REGION Network 8: Störungsgruppe 2 und Änderung ermitteln; Bits -> DB für Anzeige
         L     4;  // Interner Offset für Störungsgruppe 2
         SLD   3;  // Anzahl der Bytes für die StGrp 1
         LAR1;  // Adresse für lokale Störungen
   //
         L     4;  // Interner Offset für Störungsgruppe 2
         L     #IN_Start_Stoerungen;
         +D;
         SLD   3;  //
         LAR2;  // Adresse für Störung im DB
   //
         L     1;  // Anzahl der Störungsworte
   M004: T     #Schleifenzaehler;  // Wenn Schleifenzähler <> 0
   //
         OPN   #IN_DB_Stoerungen;  //
         L     DBW[AR2, P#0.0];  // Gespeicherte Störung mit
         L     LW[AR1, P#0.0];  // Lokale Störung       vergleichen
         <>D;  //
         T     DBW[AR2, P#0.0];  // im DB speichern und
         S     #IO_Daten_Senden;  // Sendeanforderung an PU (FB120)
         S     #IO_Stoerungsaenderung;  // Störungsanderung für Störauswertung (FB9)
         S     #IO_Stoer_Grp_2_aktiv;  // und Sammelsignal setzen
   //
         +AR1  P#2.0;
         +AR2  P#2.0;
   //
         L     #Schleifenzaehler;  // Wenn Schleifenzähler <> 0
         LOOP  M004;  // Schleife erneut durchlaufen
   //
         A     #IN_Stoer_Grp_2_von_Ext;  // Störung vom Rechner
         AN    #IN_Reset_fault_Grp;  // in die SPS einbinden
         FP    #IO_FM_Stoer_Grp_2_v_Ext;
         S     #IO_Stoerungsaenderung;
         S     #IO_Stoer_Grp_2_aktiv;
END_REGION

REGION Network 9: Störungsgruppe 3 und Änderung ermitteln; Bits -> DB für Anzeige
         L     6;  // Interner Offset für Störungsgruppe 3
         SLD   3;  // Anzahl der Bytes für die StGrp 1 +2
         LAR1;  // Adresse für lokale Störungen
   //
         L     6;  // Interner Offset für Störungsgruppe 3
         L     #IN_Start_Stoerungen;
         +D;
         SLD   3;  //
         LAR2;  // Adresse für Störung im DB
   //
         L     3;  // Anzahl der Störungsworte
   M005: T     #Schleifenzaehler;  //
   //
         OPN   #IN_DB_Stoerungen;  //
         L     DBW[AR2, P#0.0];  // Gespeicherte Störung mit
         L     LW[AR1, P#0.0];  // Lokale Störung       vergleichen
         <>D;  //
         T     DBW[AR2, P#0.0];  // im DB speichern und
         S     #IO_Daten_Senden;  // Sendeanforderung an PU (FB120)
         S     #IO_Stoerungsaenderung;  // Störungsanderung für Störauswertung (FB9)
         S     #IO_Stoer_Grp_3_aktiv;  // und Sammelsignal setzen
   //
         +AR1  P#2.0;
         +AR2  P#2.0;
   //
         L     #Schleifenzaehler;  // Wenn Schleifenzähler <> 0
         LOOP  M005;  // Schleife erneut durchlaufen
   //
         A     #IN_Stoer_Grp_3_von_Ext;  // Storung vom Rechner
         AN    #IN_Reset_fault_Grp;  // in die SPS einbinden
         FP    #IO_FM_Stoer_Grp_3_v_Ext;
         S     #IO_Stoerungsaenderung;
         S     #IO_Stoer_Grp_3_aktiv;
END_REGION

REGION Network 10: Meldungen und Änderung ermitteln; Bits -> DB für Anzeige
         L     12;  // Interner Offset für Meldungen
         SLD   3;  //
         LAR1;  // Adresse für lokale Störungen
   //
         L     12;  // Interner Offset für Meldungen
         L     #IN_Start_Stoerungen;
         +D;
         SLD   3;  //
         LAR2;  // Adresse für Störung im DB
   //
         L     2;  // Anzahl der Meldungsworte
   M007: T     #Schleifenzaehler;  //
   //
         OPN   #IN_DB_Stoerungen;  //
         L     DBW[AR2, P#0.0];  // Gespeicherte Störung mit
         L     LW[AR1, P#0.0];  // Lokale Störung       vergleichen
         <>D;  //
         T     DBW[AR2, P#0.0];  // im DB speichern und
         S     #IO_Daten_Senden;  // Sendeanforderung an PU (FB120)
   //
         +AR1  P#2.0;
         +AR2  P#2.0;
   //
         L     #Schleifenzaehler;  // Wenn Schleifenzähler <> 0
         LOOP  M007;  // Schleife erneut durchlaufen
END_REGION
END_FUNCTION

FUNCTION "FC1019_Stoerauswertung" : Void   // FC1019, STL
TITLE = Stoerungsquittierung für 1 Formträger
{ S7_Optimized_Access := 'FALSE' }
AUTHOR : KT242
VERSION : 0.1
// Die Stoerungsquittierung erfolgt in zwei SPS-Zyklen: 
// 1.: mit Reset_fault_Fkt werden die Störungsbits der einzelnen FCs zurückgesetzt
// 2.: mit Reset_fault_Grp werden die Störungsbits der FCs für die Störungsgruppen
//     zurückgesetzt. Bilden diese nun die Störungen neu, so werten sie von
//     den einzelnen FCs bereits den aktuellen Stand aus, da diese bereits einen
//     SPS-Zyklus früher bearbeitet wurden.
// 
// Das Ablöschen der Störungen in der Visualisierung wird von den einzelnen 
// Stör-FCs organisiert.
   VAR_INPUT
      IN_Stoer_Grp_1_aktiv_RT : Bool;   // Störungsmerker für eine aktive Störung der Gruppe 1 an dem Rundtisch
      IN_Stoer_Grp_2_aktiv_RT : Bool;   // Störungsmerker für eine aktive Störung der Gruppe 2 an dem Rundtisch
      IN_Stoer_Grp_3_aktiv_RT : Bool;   // Störungsmerker für eine aktive Störung der Gruppe 3 an dem Rundtisch
      IN_Taster_Quittierung : Bool;   // Eingang für einen Taster zum quittieren der Störungen
      IN_Lampentest : Bool;   // Zur Überprüfung der Anzeigen wurde ein Lampentest angewählt
      IN_Erster_SPS_Zyklus : Bool;   // Impulssignal Neusstart der Steuerung zum ablöschen der Störungen
   END_VAR
   VAR_OUTPUT
      OUT_akustische_Anzeige : Bool;   // Ausgang für eine akustische Störungsanzeige (Nur bei Neustörungen)
      OUT_optische_Anzeige : Bool;   // Ausgang für eine optische Störungsanzeige
   END_VAR
   VAR_IN_OUT
      IO_Erste_Quittierung_oK : Bool;   // Hilfsmerker zum ablöschen der akustischen Störanzeige nach Quittierung
      IO_Reset_fault_Fkt : Bool;   // Signal zum quittieren der Störungen innerhalb der einzelnen Funktionsbausteine
      IO_Reset_fault_Grp : Bool;   // Signal zum quittieren der Störungen innerhalb der Störungsbausteine
      Stoerungsaenderung : Bool;   // Feststellen einer Störungsänderung für Abarbeitung
      IO_Quit_Flanke : Bool;   // Hilkfsmerker zur Überwachung der Betätigung des Quittiertasters
   END_VAR
   VAR_TEMP
      Sammel_Stoerung : Bool;   // Zwischenmerker für die erkennung einer anliegenden Störung
      Quit_Flanke : Bool;   // Zwischenmerker als Impuls für die Störungsquittierung
      Lampe_ein : Bool;   // Zwischenmerker für die Ansteuerung der optischen Störanzeige
   END_VAR
BEGIN

REGION Network 1: Störungsquittierung für die SPS
         NOP   0;
   //
   // Über das Bit Reset_fault_Fkt werden zuerst die Störungen
   // in den Funktionen in dem sie gebildet werden abgelöscht.
   // Im nächsten SPS- Zyklus werden dann erst die Störbits
   // in den jeweiligen Störungsbausteinen abgelöscht
   //
         A     #IO_Reset_fault_Grp;  // Für den Störungsbaustein
         R     #IO_Reset_fault_Grp;
   //
         A     #IO_Reset_fault_Fkt;  // Für die einzelnen Funktionsbausteine
         S     #IO_Reset_fault_Grp;
         R     #IO_Reset_fault_Fkt;
   //
   // Bilden einer Sammelstörung
   //
         O     #IN_Stoer_Grp_1_aktiv_RT;
         O     #IN_Stoer_Grp_2_aktiv_RT;
         O     #IN_Stoer_Grp_3_aktiv_RT;
         =     #Sammel_Stoerung;
   //
   // Quittierflanke gegen Dauerbetätigung des Quittiertasters
   //
         A     #IN_Taster_Quittierung;
         FP    #IO_Quit_Flanke;
         =     #Quit_Flanke;
   //
   // Wenn keine Störung mehr ansteht oder
   // wenn eine neue Störungsänderung erfolgt,
   // wird das Bit für die erste Quittierung zurückgesetzt
   //
         O     #Stoerungsaenderung;
         ON    #Sammel_Stoerung;
         R     #IO_Erste_Quittierung_oK;
   //
   // Wenn Störungen anstehen und zum 2´ten mal quittiert
   // wird wird das Quittierbit für die einzelnen FC´s
   // gesetzt
   //
         A     #Sammel_Stoerung;
         A     #IO_Erste_Quittierung_oK;
         A     #Quit_Flanke;
         S     #IO_Reset_fault_Fkt;
   //
   // Wurde die 2´te Quittierung an die einzelnen Maschinen
   // weitergegeben wird der Merker für die 1´te Quittierung
   // zurückgesetzt
   //
         A     #IO_Reset_fault_Fkt;
         R     #IO_Erste_Quittierung_oK;
   //
   // 1´tes mal quittieren -> Hupe ausschalten
   //
         A     #Sammel_Stoerung;
         AN    #Stoerungsaenderung;
         A     #Quit_Flanke;
         AN    #IO_Reset_fault_Fkt;
         S     #IO_Erste_Quittierung_oK;
   //
   // Störlampe immer wenn eine Störung ansteht
   //
         A     #Sammel_Stoerung;
         A     "Flag_01_000_Hertz";
         =     #Lampe_ein;
         O     #Lampe_ein;
         O     #IN_Lampentest;
         =     #OUT_optische_Anzeige;
   //
   // Störhupe nur wenn die erste Quittierung noch nicht erfolgte
   //
         O     #Lampe_ein;
         O     #IN_Lampentest;
         AN    #IO_Erste_Quittierung_oK;
         AN    #IN_Lampentest;
         =     #OUT_akustische_Anzeige;
   //
   // Bilden der Quittierungsbits zum ablöschen der einzelnen
   // Störungrn innerhalb der Funktionsbausteine
   //
         AN    #Sammel_Stoerung;
         A     #Quit_Flanke;
         O     #IN_Erster_SPS_Zyklus;  // Neustart der Steuerung
         S     #IO_Reset_fault_Fkt;
   //
   // Das Bit für die Anzeige einer Stoerungsaenderung
   // aus dem Störungsbaustein (FC1) wird zurücksetzen
   //
         SET;
         R     #Stoerungsaenderung;
END_REGION
END_FUNCTION

FUNCTION "FC1021_TT_Operation_mode" : Void   // FC1021, STL
TITLE = Betriebsarten der Anlage
{ S7_Optimized_Access := 'TRUE' }
VERSION : 0.1
   VAR_TEMP
      FRG_Start_Produktion : Bool;
      FRG_Produktion : Bool;
      FRG_Stop : Bool;
      Stopptaster : Bool;
      STG_GRP_2 : Bool;
      Temp_Auto_Stop_ok : Bool;
      Hupe_Anfahrwarnung : Bool;
      Anf_Stop : Bool;
   END_VAR
BEGIN

REGION Network 1
         A     "AS_turn_table";
         =     #Temp_Auto_Stop_ok;
         NOT;
         =     "DB1010_TT_Fault".AS.AS_Activ;
   //      =     "TT_H_AS"
END_REGION

REGION Network 2: Freigabesignale Produktion Starten bilden
         A     "DB1001_TT_State".BA_Anlage.Automatik_Stop_ok;
         A     "DB1001_TT_State".IPOS.Status.IPOS_referenziert;
         AN    "DB1001_TT_State".Bits.Stop_fuer_WW;
         AN    "DB1031_AddStatus".SaftyDevice[1].OpeningEnabled;
         AN    "DB1031_AddStatus".SaftyDevice[2].OpeningEnabled;
         AN    "DB1031_AddStatus".SaftyDevice[3].OpeningEnabled;
         AN    "DB1031_AddStatus".SaftyDevice[4].OpeningEnabled;
         =     #FRG_Start_Produktion;
END_REGION

REGION Network 3: Freigabesignale Produktionsbetrieb bilden
         A     "DB1001_TT_State".BA_Anlage.Start_Produktion;
         A     "DB1001_TT_State".IPOS.Status.RT_in_Position;
         =     #FRG_Produktion;
END_REGION

REGION Network 4: Freigabesignale Produktion Stoppen bilden
         A     "DB1001_TT_State".IPOS.Status.Stoppen_erkannt;
         A     "DB1001_TT_State".IPOS.Status.RT_in_Position;
         AN    "DB005_RS<->Extern".MC_Interface[1].Data_from_MC.Shot_preperation;
         =     #FRG_Stop;
END_REGION

REGION Network 5: Signal zum Stoppen bilden
         A     "Button_stop_cycle";
         AN    "DB1001_TT_State".Bits.Stop_fuer_WW;
         AN    "DB1001_TT_State".Bits.Stop_fuer_Teachen;
         AN    "DB1001_TT_State".Bits.StopAfterEmpty;
         A     "DB1001_TT_State".BA_Anlage.Automatik;
         =     #Stopptaster;
END_REGION

REGION Network 6: Bei Leerfahren der Anlage Störgruppe 2 ausblenden
         A     "DB1011_TT_Fault".STG2_RT;
         =     #STG_GRP_2;
END_REGION

REGION Network 7: Stoppen angefordert
         O     "DB1001_TT_State".Bits.Stop_fuer_WW;
         O     "DB1001_TT_State".Bits.Stop_fuer_Teachen;
         =     #Anf_Stop;
END_REGION

REGION Network 8: Funktion für Betriebsart
         CALL  "FC1022_TT_OM"
         ( IN_Steuerpannung        := "Controlvoltage_okay",
           IN_SS_Auto              := "Switch_automatic_mode",
           IN_SS_Hand              := "Switch_manual_mode",
           IN_Referenzieren        := "Button_reference_TT",
           IN_Automatik_Stop_ok    := #Temp_Auto_Stop_ok,
           IN_T_Start              := "Button_start_cycle",
           IN_T_Stop               := #Stopptaster,
           IN_Lampentest           := FALSE,
           IN_Werkzeugwechsel      := #Anf_Stop,
           IN_Freigabe_Start       := #FRG_Start_Produktion,
           IN_Freigabe_Produktion  := #FRG_Produktion,
           IN_Freigabe_Stop        := #FRG_Stop,
           IN_Stoerung_Gruppe_1    := "DB1011_TT_Fault".STG1_RT,
           IN_Stoerung_Gruppe_2    := #STG_GRP_2,
           IN_DW_Maxzeit_Prod_ein  := S5T#10S,
           IN_DW_Maxzeit_Prod_aus  := S5T#30S,
           IN_DW_Zeit_Startwarnung := "DB1049_TT_Value".Vorwarnzeit,
           IN_Betriebsart_Timer    := "TMTT_OPMode",
           IN_Anfahr_Timer         := "TMTT_StartProduction",
           IN_Produktions_Timer    := "TMTT_Production",
           Out_Anfahrwarnung       := #Hupe_Anfahrwarnung,
           IO_Status               := "DB1001_TT_State".BA_Anlage
         );
   //-----
END_REGION

REGION Network 9: Anzeige der Betriebsart der Anlage
         A     "DB1001_TT_State".BA_Anlage.Start_Produktion;
         A     "Flag_01_000_Hertz";
         O;
         A     "DB1001_TT_State".BA_Anlage.Produktion;
         A     "DB1001_TT_State".BA_Anlage.Stop_angefordert;
         A     "Flag_01_000_Hertz";
         O;
         A     "DB1001_TT_State".BA_Anlage.Produktion;
         AN    "DB1001_TT_State".BA_Anlage.Stop_angefordert;
         O     "DB1001_TT_State".BA_Anlage.Lampentest;
         =     "LED_start_cycle";
END_REGION

REGION Network 10: Leerfahren der Anlage ist beendet
   //      U     "T_Leerfahren_RT_1"
   //      FP    "FHM_RT_Leerfahren_RT1"
   //      =     "HM_RT_Leerfahren_RT1"
   //
   //      X     "HM_RT_Leerfahren_RT1"
   //      X     "DB005_RS<->Extern".Status_RT_1.S_RT_Leerfahren
   //      =     "DB005_RS<->Extern".Status_RT_1.S_RT_Leerfahren
   //
   //      U     #Starttaster
   //      R     "DB005_RS<->Extern".Status_RT_1.S_RT_Leerfahren
   // //
   //       U(
   //       O     "DB201_RT1_Segment_1".Status_FT.FT_aktuell.Status.FT_gesperrt
   //       O     "DB201_RT1_Segment_1".Status_FT.FT_aktuell.Status.FT_in_Abwahlposition
   //       )
   //       U(
   //       O     "DB202_RT1_Segment_2".Status_FT.FT_aktuell.Status.FT_gesperrt
   //       O     "DB202_RT1_Segment_2".Status_FT.FT_aktuell.Status.FT_in_Abwahlposition
   //       )
   //       U(
   //       O     "DB203_RT1_Segment_3".Status_FT.FT_aktuell.Status.FT_gesperrt
   //       O     "DB203_RT1_Segment_3".Status_FT.FT_aktuell.Status.FT_in_Abwahlposition
   //       )
   //       U(
   //       O     "DB204_RT1_Segment_4".Status_FT.FT_aktuell.Status.FT_gesperrt
   //       O     "DB204_RT1_Segment_4".Status_FT.FT_aktuell.Status.FT_in_Abwahlposition
   //       )
   //       U(
   //       O     "DB205_RT1_Segment_5".Status_FT.FT_aktuell.Status.FT_gesperrt
   //       O     "DB205_RT1_Segment_5".Status_FT.FT_aktuell.Status.FT_in_Abwahlposition
   //       )
   //       U(
   //       O     "DB206_RT1_Segment_6".Status_FT.FT_aktuell.Status.FT_gesperrt
   //       O     "DB206_RT1_Segment_6".Status_FT.FT_aktuell.Status.FT_in_Abwahlposition
   //       )
   //       U(
   //       O     "DB207_RT1_Segment_7".Status_FT.FT_aktuell.Status.FT_gesperrt
   //       O     "DB207_RT1_Segment_7".Status_FT.FT_aktuell.Status.FT_in_Abwahlposition
   //       )
   //       U(
   //       O     "DB208_RT1_Segment_8".Status_FT.FT_aktuell.Status.FT_gesperrt
   //       O     "DB208_RT1_Segment_8".Status_FT.FT_aktuell.Status.FT_in_Abwahlposition
   //       )
   //       U(
   //       O     "DB209_RT1_Segment_9".Status_FT.FT_aktuell.Status.FT_gesperrt
   //       O     "DB209_RT1_Segment_9".Status_FT.FT_aktuell.Status.FT_in_Abwahlposition
   //       )
   //       U(
   //       O     "DB210_RT1_Segment_10".Status_FT.FT_aktuell.Status.FT_gesperrt
   //       O     "DB210_RT1_Segment_10".Status_FT.FT_aktuell.Status.FT_in_Abwahlposition
   //       )
   //       U(
   //       O     "DB211_RT1_Segment_11".Status_FT.FT_aktuell.Status.FT_gesperrt
   //       O     "DB211_RT1_Segment_11".Status_FT.FT_aktuell.Status.FT_in_Abwahlposition
   //       )
   //       U(
   //       O     "DB212_RT1_Segment_12".Status_FT.FT_aktuell.Status.FT_gesperrt
   //       O     "DB212_RT1_Segment_12".Status_FT.FT_aktuell.Status.FT_in_Abwahlposition
   //       )
   //       U(
   //       O     "DB213_RT1_Segment_13".Status_FT.FT_aktuell.Status.FT_gesperrt
   //       O     "DB213_RT1_Segment_13".Status_FT.FT_aktuell.Status.FT_in_Abwahlposition
   //       )
   //       U(
   //       O     "DB214_RT1_Segment_14".Status_FT.FT_aktuell.Status.FT_gesperrt
   //       O     "DB214_RT1_Segment_14".Status_FT.FT_aktuell.Status.FT_in_Abwahlposition
   //       )
   //       U(
   //       O     "DB215_RT1_Segment_15".Status_FT.FT_aktuell.Status.FT_gesperrt
   //       O     "DB215_RT1_Segment_15".Status_FT.FT_aktuell.Status.FT_in_Abwahlposition
   //       )
   //       U(
   //       O     "DB216_RT1_Segment_16".Status_FT.FT_aktuell.Status.FT_gesperrt
   //       O     "DB216_RT1_Segment_16".Status_FT.FT_aktuell.Status.FT_in_Abwahlposition
   //       )
   //       U(
   //       O     "DB217_RT1_Segment_17".Status_FT.FT_aktuell.Status.FT_gesperrt
   //       O     "DB217_RT1_Segment_17".Status_FT.FT_aktuell.Status.FT_in_Abwahlposition
   //       )
   //       U(
   //       O     "DB218_RT1_Segment_18".Status_FT.FT_aktuell.Status.FT_gesperrt
   //       O     "DB218_RT1_Segment_18".Status_FT.FT_aktuell.Status.FT_in_Abwahlposition
   //       )
   //       U(
   //       O     "DB219_RT1_Segment_19".Status_FT.FT_aktuell.Status.FT_gesperrt
   //       O     "DB219_RT1_Segment_19".Status_FT.FT_aktuell.Status.FT_in_Abwahlposition
   //       )
   //       U(
   //       O     "DB220_RT1_Segment_20".Status_FT.FT_aktuell.Status.FT_gesperrt
   //       O     "DB220_RT1_Segment_20".Status_FT.FT_aktuell.Status.FT_in_Abwahlposition
   //       )
   //       =     "DB005_RS<->Extern".Status_RT_1.RT_ist_leergefahren
   // //
   //       U     "DB005_RS<->Extern".Status_RT_1.S_RT_Leerfahren
   //       UN    "DB005_RS<->Extern".Status_RT_1.RT_ist_leergefahren
   //       U     "Merker_01_000_Hertz"
   //       O(
   //       U     "DB005_RS<->Extern".Status_RT_1.RT_ist_leergefahren
   //       U     "DB005_RS<->Extern".Status_RT_1.S_RT_Leerfahren
   //       )
   //       O     "DB151_Rundtisch_1".BA_Anlage.Lampentest
   //       =     "H_Leerfahren_RT_1"
END_REGION
END_FUNCTION

FUNCTION "FC1022_TT_OM" : Void   // FC1022, STL
TITLE = Betriebsarten für die Anlage
{ S7_Optimized_Access := 'FALSE' }
AUTHOR : KT242
VERSION : 0.1
// Die Verwaltung der Betriebsarten geschieht wie folgt: 
// Die Betriebsarten hängen nur von der Stellung des Betriebsartenwahlschalters 
// ab, wie man es z.B. auch bei Robotern gewohnt ist. Das Bit "gültig" wurde in 
// "aktiv" geändert und zeigt zusätzlich, dass Steuerspannung und Schutztüren 
// o.k. sind.
// Referenzpunktfahren ist keine Betriebsart sondern ein zusätzliches Bit in 
// Betriebsart Hand.
// Automatikbetrieb hängt nicht davon ab, ob es möglich ist, die Anlage zu 
// bewegen. 
// Aggregate, die für den Automatikbetrieb nötig sind, sollten schon eingeschaltet 
// werden, wenn Betriebsart Automatik anliegt und Steuerspannung und NOTHALT o.k.
// sind.
   VAR_INPUT
      IN_Steuerpannung : Bool;   // Signal Steuerspannung Eingeschaltet und Not- Aus entriegelt
      IN_SS_Auto : Bool;   // Eingang Betriebsartenwahlschalter steht auf Automatik- Betrieb
      IN_SS_Hand : Bool;   // Eingang Betriebsartenwahlschalter steht auf Hand- Betrieb
      IN_Referenzieren : Bool;   // Eingang Taster für Referenzpunktfahrt
      IN_Automatik_Stop_ok : Bool;   // Eingang das die Sicherheitseinrichtungen quittiert sind
      IN_T_Start : Bool;   // Eingang für den Taster zum Starten des Rundtisches
      IN_T_Stop : Bool;   // Eingang für den Taster zum Stoppen des Rundtisches
      IN_Lampentest : Bool;   // Eingang für eine Funktionsüberprüfung der Lampenansteuerungen
      IN_Werkzeugwechsel : Bool;   // Signal das ein Werkzeugwechsel vorgewählt wurde
      IN_Freigabe_Start : Bool;   // Signal für die Freigabe zum Starten des Rundtisches
      IN_Freigabe_Produktion : Bool;   // Signal für die Freigabe des Produktionsbetriebes des Rundtisches
      IN_Freigabe_Stop : Bool;   // Signal für die Freigabe zum Stoppen des Rundtisches
      IN_Stoerung_Gruppe_1 : Bool;   // Eine Störung der Gruppe 1 steht an und wurde noch nicht quittiert
      IN_Stoerung_Gruppe_2 : Bool;   // Eine Störung der Gruppe 2 steht an und wurde noch nicht quittiert
      IN_DW_Maxzeit_Prod_ein : S5Time;   // Zeit in der die Produktion nach dem Starten freigegeben sein muß
      IN_DW_Maxzeit_Prod_aus : S5Time;   // Verzögerungszeit zum Stoppen des Produktionsbetriebes
      IN_DW_Zeit_Startwarnung : S5Time;   // Ansteuerungsdauer für eine Anfahrwarnung
      IN_Betriebsart_Timer : Timer;   // Timer für die Betriebsartenumschaltung
      IN_Anfahr_Timer : Timer;   // Timer für die Anfahrwarnung der Anlage
      IN_Produktions_Timer : Timer;   // Timer für die Produktions Start- und Abschaltung
   END_VAR
   VAR_OUTPUT
      Out_Anfahrwarnung : Bool;   // Ansteuerung einer Anfahrwarnung
   END_VAR
   VAR_IN_OUT
      IO_Status : "UDT_RT_Betriebsart";   // Speichern der Betriebsarten- Zustände für das Programm
   END_VAR
   VAR_TEMP
      Temp_IO_Status : "UDT_RT_Betriebsart";   // Temporärer Betriebsarten- Status für die interne Bearbeitung des Bausteins
      ERROR_CODE : Int;   // Störungszustand der Systemfunktion "BLKMOV" Blockmove
      Anyzeiger : ANY;   // Zeiger zum Kopieren der Bereiche "IO_Status" und "Temp_IO_Status"
      Ohne_Anfahrwarnung : Bool;   // Hilfsmerker das keine Anfahrwarnung benötigt wird
      Temp_Imp_Anfahrwarn_End : Bool;   // Impulsmerker das die Anfahrwarnung gerade beendet wurde
   END_VAR
BEGIN

REGION Network 1: Gesicherte Daten einbinden
         LAR1;
         L;
         LAR2;
   //
         L     W#16#1002;  // Bytes
         T     W[AR1, P#0.0];
         L     2;  // Anzahl Bytes
         T     W[AR1, P#2.0];
         L     W[AR2, P#0.0];  // Baustein Nr.
         T     W[AR1, P#4.0];
         L     D[AR2, P#2.0];  // Datenanfang
         T     D[AR1, P#6.0];
   //
         CALL  BLKMOV
         ( SRCBLK  := #Anyzeiger,
           RET_VAL := #ERROR_CODE,
           DSTBLK  := #Temp_IO_Status
         );
   //
END_REGION

REGION Network 2: Automatik- Stop
         A     #IN_Automatik_Stop_ok;
         =     #Temp_IO_Status.Automatik_Stop_ok;
END_REGION

REGION Network 3: Steuerspannung vorhanden
         A     #IO_Status.Steuerspannung_ein;
         JC    Spg;
   //
         A     #IN_Steuerpannung;
         L     S5T#1S;
         SD    #IN_Betriebsart_Timer;
         A     #IN_Betriebsart_Timer;
         =     #Temp_IO_Status.Steuerspannung_ein;
         JU    BA;
   //
   Spg:  A     #IN_Steuerpannung;
         =     #Temp_IO_Status.Steuerspannung_ein;
END_REGION

REGION Network 4: Wechsel der Betriebsart
         O(;
         AN    #IN_SS_Hand;
         A     #Temp_IO_Status.Hand;
         );
         O(;
         AN    #IN_SS_Auto;
         A     #Temp_IO_Status.Automatik;
         );
         L     S5T#500MS;
         SE    #IN_Betriebsart_Timer;
         A     #IN_Betriebsart_Timer;
         JC    GOON;
END_REGION

REGION Network 5: Betriebsartenschalter-Auswertung
   BA:   A     #IN_SS_Hand;
         AN    #IN_SS_Auto;
         =     #Temp_IO_Status.Hand;
   //
         AN    #IN_SS_Hand;
         A     #IN_SS_Auto;
         =     #Temp_IO_Status.Automatik;
   //
   GOON: A     #IN_Lampentest;
         =     #Temp_IO_Status.Lampentest;
   //
         O     #Temp_IO_Status.Hand;
         O     #Temp_IO_Status.Automatik;
         =     #Temp_IO_Status.Gueltig;
   //
         O     #Temp_IO_Status.Hand;
         O     #Temp_IO_Status.Automatik;
         A     #Temp_IO_Status.Steuerspannung_ein;
         A     #Temp_IO_Status.Automatik_Stop_ok;
         =     #Temp_IO_Status.Aktiv;
   //
         A     #Temp_IO_Status.Hand;
         A     #IN_Referenzieren;
         =     #Temp_IO_Status.Referenzieren;
END_REGION

REGION Network 6: Ausgabe eines Startsignales vor Ansteuerung der Anlage
         L     #IN_DW_Zeit_Startwarnung;
         L     0;
         ==D;
         =     #Ohne_Anfahrwarnung;
   //
         L     #IN_DW_Zeit_Startwarnung;
         A     #IN_Freigabe_Start;
         A     #IN_T_Start;
         A     #IN_T_Stop;
         A     #Temp_IO_Status.Automatik;
         AN    #IN_Stoerung_Gruppe_1;
         AN    #IN_Stoerung_Gruppe_2;
         AN    #Temp_IO_Status.Produktion;
         AN    #Temp_IO_Status.Start_Produktion;
         SE    #IN_Anfahr_Timer;
   //
         A     #IN_Anfahr_Timer;
         =     #Temp_IO_Status.Anfahrwarnung;
   //
         A     #Temp_IO_Status.Anfahrwarnung;
         =     #Out_Anfahrwarnung;
   //
         AN    #Temp_IO_Status.Anfahrwarnung;
         FP    #Temp_IO_Status.FHM_Anfahrwarnung;
         =     #Temp_Imp_Anfahrwarn_End;
END_REGION

REGION Network 7: Bit für Start Produktion
         L     #IN_DW_Maxzeit_Prod_ein;
         A     #IN_T_Start;
         A     #Ohne_Anfahrwarnung;
         O     #Temp_Imp_Anfahrwarn_End;
         A     #IN_Freigabe_Start;
         AN    #Temp_IO_Status.Produktion;
         AN    #Temp_IO_Status.Start_Produktion;
         S     #Temp_IO_Status.Start_Produktion;
         SE    #IN_Produktions_Timer;
   //
         ON    #IN_Produktions_Timer;
         ON    #Temp_IO_Status.Aktiv;
         ON    #Temp_IO_Status.Automatik;
         O     #IN_Stoerung_Gruppe_1;
         O     #IN_Stoerung_Gruppe_2;
         ON    #IN_T_Stop;
         O     #IN_Werkzeugwechsel;
         ON    #Temp_IO_Status.Automatik_Stop_ok;
         R     #Temp_IO_Status.Start_Produktion;
END_REGION

REGION Network 8: Bit für Produktion
         A     #Temp_IO_Status.Start_Produktion;
         A     #IN_Freigabe_Produktion;
         AN    #IN_Anfahr_Timer;
         S     #Temp_IO_Status.Produktion;
         R     #Temp_IO_Status.Start_Produktion;
   //
         L     #IN_DW_Maxzeit_Prod_aus;
         ON    #IN_T_Stop;
         O     #IN_Werkzeugwechsel;
         O     #IN_Stoerung_Gruppe_2;
         A     #Temp_IO_Status.Produktion;
         AN    #Temp_IO_Status.Stop_angefordert;
         S     #Temp_IO_Status.Stop_angefordert;
         SE    #IN_Produktions_Timer;
   //
         A     #Temp_IO_Status.Produktion;
         A     #IN_T_Start;
         AN    #IN_Werkzeugwechsel;
         R     #Temp_IO_Status.Stop_angefordert;
   //
         A     #Temp_IO_Status.Produktion;
         A     #Temp_IO_Status.Stop_angefordert;
         AN    #IN_Produktions_Timer;
         O;
         A     #Temp_IO_Status.Produktion;
         A     #Temp_IO_Status.Stop_angefordert;
         A     #IN_Freigabe_Stop;
         O     #IN_Stoerung_Gruppe_1;
         ON    #Temp_IO_Status.Automatik;
         ON    #Temp_IO_Status.Automatik_Stop_ok;
         ON    #Temp_IO_Status.Aktiv;
         R     #Temp_IO_Status.Produktion;
         R     #Temp_IO_Status.Stop_angefordert;
END_REGION

REGION Network 9: Daten sichern
         CALL  BLKMOV
         ( SRCBLK  := #Temp_IO_Status,
           RET_VAL := #ERROR_CODE,
           DSTBLK  := #Anyzeiger
         );
   //
END_REGION
END_FUNCTION

FUNCTION "FC1031_AdditionalDevice" : Void   // FC1031, STL
{ S7_Optimized_Access := 'TRUE' }
VERSION : 0.1
   VAR_TEMP
      Release_door : Bool;
      dummy : Bool;
   END_VAR
BEGIN

REGION Network 1: Safety door tool change
   //      UN    "DB1001_TT_State".BA_Anlage.Start_Produktion
   //      UN    "DB1001_TT_State".BA_Anlage.Produktion
   //      =     #Release_door
   //
   //      CALL  "FC1033_SafetyDevice"
   //         IN_With_Safety_door :=TRUE //"Settings_MCx".MC_settings.MCwithSafetydoor
   //         IN_EnableDoorOpen   :=#Release_door
   //         IN_SelectDoorOpen   :="Select_door_tool_change"
   //         IN_AS_Door          :="AS_door_tool_change"
   //         IN_QuitDoorOpen     :="Quit_door_tool_change"
   //         IN_OMLampTest       :="DB1001_TT_State".BA_Anlage.Lampentest
   //         IN_Delay_QuitDoor   :="TM_QuitDoor_MC1"
   //         OUT_V_DoorOpen      :="Release_door_tool_change"
   //         OUT_H_DoorOpen      :="Selected_door_tool_change"
   //         StatusSafetyDevice  :="DB1031_AddStatus".SaftyDevice[1]
END_REGION

REGION Network 2: Safety door robot
   //      UN    "DB1001_TT_State".BA_Anlage.Start_Produktion
   //      UN    "DB1001_TT_State".BA_Anlage.Produktion
   //      =     #Release_door
   //
   //      CALL  "FC1033_SafetyDevice"
   //         IN_With_Safety_door :=TRUE //"Settings_MCx".MC_settings.MCwithSafetydoor
   //         IN_EnableDoorOpen   :=#Release_door
   //         IN_SelectDoorOpen   :="Select_door_robot"
   //         IN_AS_Door          :="AS_door_robot"
   //         IN_QuitDoorOpen     :="Quit_door_robot"
   //         IN_OMLampTest       :="DB1001_TT_State".BA_Anlage.Lampentest
   //         IN_Delay_QuitDoor   :="TM_QuitDoor_MC1"
   //         OUT_V_DoorOpen      :="Release_door_robot"
   //         OUT_H_DoorOpen      :="Selected_door_robot"
   //         StatusSafetyDevice  :="DB1031_AddStatus".SaftyDevice[2]
END_REGION

REGION Network 3: Safety door test shot
END_REGION

REGION Network 4: Safety door turn table
   //      UN    "DB1001_TT_State".BA_Anlage.Start_Produktion
   //      UN    "DB1001_TT_State".BA_Anlage.Produktion
   //      =     #Release_door
   //
   //      CALL  "FC1033_SafetyDevice"
   //         IN_With_Safety_door :=TRUE //"Settings_MCx".MC_settings.MCwithSafetydoor
   //         IN_EnableDoorOpen   :=#Release_door
   //         IN_SelectDoorOpen   :="Select_door_TT"
   //         IN_AS_Door          :="AS_door_TT"
   //         IN_QuitDoorOpen     :="Quit_door_TT"
   //         IN_OMLampTest       :="DB1001_TT_State".BA_Anlage.Lampentest
   //         IN_Delay_QuitDoor   :="TM_QuitDoor_MC1"
   //         OUT_V_DoorOpen      :="Release_door_TT"
   //         OUT_H_DoorOpen      :="Selected_door_TT"
   //         StatusSafetyDevice  :="DB1031_AddStatus".SaftyDevice[3]

   //
END_REGION
END_FUNCTION

FUNCTION "FC1032_PneuZylindermSH" : Void   // FC1032, STL
TITLE = Pneumatischer Zylinder mit Selbsthaltung
{ S7_Optimized_Access := 'FALSE' }
VERSION : 0.1
   VAR_INPUT
      BA_Auto : Bool;   // Betriebsart Automatik
      BA_Hand : Bool;   // Tippbetrieb
      Anf_GS : Bool;   // Anforderung Grundstellung Automatik
      Anf_AS : Bool;   // Anforderung Arbeitsstellung Automatik
      T_GS : Bool;   // Taste Grundstellung (Tippbetrieb)
      T_AS : Bool;   // Taste Arbeitsstellung (Tippbetrieb)
      Frg_GS : Bool;   // Bewegungsbedingungen für Grundstellungsfahrt erfüllt
      Frg_AS : Bool;   // Bewegungsbedingungen für Arbeitstellungsfahrt erfüllt
      INI_GS : Bool;   // Sensorik Zylinder befindet sich in Grundstellung
      INI_AS : Bool;   // Sensorik Zylinder befindet sich in Arbeitsstellung
      P_GS : Bool;   // Druckschalter Grundstellung
      P_AS : Bool;   // Druckschalter Arbeitsstellung
      IN_Reset_fault_Fkt : Bool;   // Signal to acknowledge faults in functionblock
      Laufzeit : S5Time;   // Laufzeit für Laufzeitüberwachung
      TM_Laufzeit : Timer;   // Timer zur Laufzeitüberwachung
   END_VAR
   VAR_OUTPUT
      H_GS : Bool;   // Anzeige Grundstellung
      H_AS : Bool;   // Anzeige Arbeitsstellung
      OUT_V_GS : Bool;   // Ventil zur Ansteuerung der Grundstellung
      OUT_V_AS : Bool;   // Ventil zur Ansteuerung der Arbeitsstellung
   END_VAR
   VAR_IN_OUT
      IO_Stg_INI : Bool;   // Sensorstörung
      IO_Stg_Laufzeit : Bool;   // Laufzeitstörung
      IO_NewFault : Bool;
      IO_FaultLevel_1 : Bool;
   END_VAR
   VAR_TEMP
      Temp_V_GS : Bool;
      Temp_V_AS : Bool;
   END_VAR
BEGIN

REGION Network 1: Ausgänge Rücksetzen
         CLR;
         =     #Temp_V_GS;
         =     #Temp_V_AS;
END_REGION

REGION Network 2: Störungen zurücksetzen
         A     #IN_Reset_fault_Fkt;
         R     #IO_Stg_INI;
         R     #IO_Stg_Laufzeit;
END_REGION

REGION Network 3: Tippbetrieb
         A     #BA_Hand;
         JCN   nHnd;

   // Arbeitsstellung
         A     #T_AS;
         A     #Frg_AS;
         O(;
         A     #INI_AS;
         A     #P_AS;
         AN(;
         A     #T_GS;
         A     #Frg_GS;
         );
         );
         =     #Temp_V_AS;

   // Grundstellung
         A     #T_GS;
         A     #Frg_GS;
         O(;
         A     #INI_GS;
         A     #P_GS;
         AN(;
         A     #T_AS;
         A     #Frg_AS;
         );
         );
         =     #Temp_V_GS;

   nHnd: NOP   0;
END_REGION

REGION Network 4: Automatik
         A     #BA_Auto;
         JCN   nAut;

   // Arbeitsstellung
         A     #Anf_AS;
         A     #Frg_AS;
         O(;
         A     #INI_AS;
         A     #P_AS;
         AN(;
         A     #Anf_GS;
         A     #Frg_GS;
         );
         );
         =     #Temp_V_AS;

   // Grundstellung
         A     #Anf_GS;
         A     #Frg_GS;
         O(;
         A     #INI_GS;
         A     #P_GS;
         AN(;
         A     #Anf_AS;
         A     #Frg_AS;
         );
         );
         =     #Temp_V_GS;

   nAut: NOP   0;
END_REGION

REGION Network 5: Anzeigen

         A     #Temp_V_GS;
         =     #OUT_V_GS;
         A     #Temp_V_AS;
         =     #OUT_V_AS;

         ON    #INI_GS;
         ON    #P_GS;
         A     #Temp_V_GS;
         A     "Flag_01_250_Hertz";
         O(;
         A     #INI_GS;
         A     #P_GS;
         );
         =     #H_GS;

         ON    #INI_AS;
         ON    #P_AS;
         A     #Temp_V_AS;
         A     "Flag_01_250_Hertz";
         O(;
         A     #INI_AS;
         A     #P_AS;
         );
         =     #H_AS;
END_REGION

REGION Network 6: Störungen
   //  Sensorstörung
         A     #INI_GS;
         A     #INI_AS;
         AN    #IO_Stg_INI;
         S     #IO_NewFault;
         S     #IO_Stg_INI;

   //  Laufzeitstörung
         A(;

         O(;
         X     #Temp_V_GS;
         X(;
         A     #INI_GS;
         A     #P_GS;
         );
         );

         O(;
         X     #Temp_V_AS;
         X(;
         A     #INI_AS;
         A     #P_AS;
         );
         );
         );

         A(;
         O     #BA_Hand;
         O     #BA_Auto;
         );

         L     #Laufzeit;
         SD    #TM_Laufzeit;

         A     #TM_Laufzeit;
         AN    #IO_Stg_Laufzeit;
         S     #IO_NewFault;
         S     #IO_Stg_Laufzeit;
END_REGION
END_FUNCTION

FUNCTION "FC1033_SafetyDevice" : Void   // FC1033, STL
{ S7_Optimized_Access := 'FALSE' }
VERSION : 0.1
   VAR_INPUT
      IN_With_Safety_door : Bool;   // Input if safety door is available
      IN_EnableDoorOpen : Bool;   // Enable signal for the release to open the door
      IN_SelectDoorOpen : Bool;   // Input for the selection to open the door
      IN_AS_Door : Bool;   // Input from the saftey that the door is open
      IN_QuitDoorOpen : Bool;   // Input to reset the door clamping
      IN_OMLampTest : Bool;   // Operation mode for lamp test is selected
      IN_Delay_QuitDoor : Timer;
   END_VAR
   VAR_OUTPUT
      OUT_V_DoorOpen : Bool;   // Output valve to clamp the door
      OUT_H_DoorOpen : Bool;   // Output for the lamp
   END_VAR
   VAR_IN_OUT
      StatusSafetyDevice : "UDT_SafetyDevice";
   END_VAR
BEGIN

REGION Network 1: If deselect jump to delete
         A     #IN_With_Safety_door;
         JCN   delete;
END_REGION

REGION Network 2: Edge of the button to select opening of the safety device
   // Switch off delay for PILZ switch

         A     #IN_QuitDoorOpen;
         L     s5t#1s;
         SF    #IN_Delay_QuitDoor;
   //----
         A     #IN_SelectDoorOpen;
         FN    #StatusSafetyDevice.HFEdgeButton;
         =     #StatusSafetyDevice.EdgeButton;
   //----
         A     #IN_AS_Door;
         FP    #StatusSafetyDevice.HFEdgeASReset;
         =     #StatusSafetyDevice.EdgeASReset;
   //----
         X     #StatusSafetyDevice.EdgeButton;
         X     #StatusSafetyDevice.OpeningSelected;
         O     #StatusSafetyDevice.HFforMESAutomaticStop;
         AN    #StatusSafetyDevice.EdgeASReset;
         AN    #IN_Delay_QuitDoor;
         =     #StatusSafetyDevice.OpeningSelected;
   //----
         A     #StatusSafetyDevice.OpeningSelected;
         A     #IN_EnableDoorOpen;
   //      ON    #IN_Delay_QuitDoor
         =     #StatusSafetyDevice.OpeningEnabled;
         NOT;
         =     #OUT_V_DoorOpen;
   //----
         O     #StatusSafetyDevice.OpeningEnabled;
         O(;
         A     #StatusSafetyDevice.OpeningSelected;
         A     "Flag_01_000_Hertz";
         );
         ON    #IN_AS_Door;
         O     #IN_OMLampTest;
         =     #OUT_H_DoorOpen;
   //----
         A     #StatusSafetyDevice.OpeningSelected;
         =     #StatusSafetyDevice.HFforMESSelected;
   //----
         AN    #IN_AS_Door;
         =     #StatusSafetyDevice.HFforMESAutomaticStop;
         R     #StatusSafetyDevice.HFforMESSelected;
   //---
         A     #StatusSafetyDevice.HFforMESSelected;
         =     #StatusSafetyDevice.Msg_Selected;
         A     #StatusSafetyDevice.HFforMESAutomaticStop;
         =     #StatusSafetyDevice.Msg_AS_active;
   //---
         BEU;
END_REGION

REGION Network 3: Delete
   delete:SET;
         R     #StatusSafetyDevice.Msg_Selected;
         R     #StatusSafetyDevice.Msg_AS_active;
         R     #OUT_H_DoorOpen;
         R     #OUT_V_DoorOpen;
END_REGION
END_FUNCTION

FUNCTION "FC1040_TT_Movement" : Void   // FC1040, STL
TITLE = Ansteuern der Anlage
{ S7_Optimized_Access := 'TRUE' }
VERSION : 0.1
   VAR_TEMP
      Temp_Segmentinis : DWord;   // Hilfsmerker für die Positionserkennung über die Hardwareabschaltung im Zentrum
      Temp_Rampe_Plus : Int;   // Hilfswort für die Beschleunigung des Rundtisches
      Temp_Rampe_Minus : Int;   // Hilfswort für die Verzögerung des Rundtisches
      Temp_Speed_Hand : Int;   // Hilfswort für die Geschwindigkeit im Handbetrieb
      Temp_Speed_Automatik : Int;   // Hilfswort für die Geschwindigkeit im Automatikbetrieb
      Temp_Offset_Position : Int;   // Hilfswort für den negativen Offset bei einer Positionierung im kont. Betrieb
      Temp_AmoutOfSegments : Int;   // Help word to define the amount of segments
      Temp_Drehsperre : Bool;   // Hilfsmerker für die generelle Freigabe dere Anlage
      Temp_Taktfreigabe : Bool;   // Hilfsmerker für das Takten der Anlage
      Temp_Drehfreigabe : Bool;   // Hilfsmerker für die Freigabe zum Ansteuern der Anlage
      Temp_RT_in_Position : Bool;   // Hilfsmerker für die Umschaltung der Segmentpositionen
      Temp_GenauhalteSignal : Bool;   // Hilfsmerker für die Ermittlung des Genauhaltes
      Temp_AnfahrWarnung : Bool;   // Hilfsmerker für die Huppe als Anfahr Warnung
      Temp_AnfahrWarnung_1 : Bool;   // Hilfsmerker für die Huppe als Anfahr Warnung
   END_VAR
BEGIN

REGION Network 1: Amount of Segments
         L     4;
         T     #Temp_AmoutOfSegments;
END_REGION

REGION Network 2: Drehsperren auswerten
         A     "DB1001_TT_State".BA_Anlage.Automatik_Stop_ok;
   //      UN    "DB009_Faults".Faults_FKT_Grp_1_M1
         =     #Temp_Drehfreigabe;
         NOT;
         =     #Temp_Drehsperre;
END_REGION

REGION Network 3: Taktzeitverlängerung // Anlage anhalten
         A     "Button_extend_cycle";
         FP    "FHM_Takt_Verz_RT1";
         =     "HM_FP_Takt_Verz_RT1";

         A     "HM_FP_Takt_Verz_RT1";
         AN    "DB1001_TT_State".Bits.Taktdehnung;
         S     "DB1001_TT_State".Bits.Taktdehnung;
         JC    VERZ;

         A     "HM_FP_Takt_Verz_RT1";
         A     "DB1001_TT_State".Bits.Taktdehnung;
         R     "DB1001_TT_State".Bits.Taktdehnung;

   VERZ: NOP   0;
         ON    "DB1001_TT_State".BA_Anlage.Produktion;
         R     "DB1001_TT_State".Bits.Taktdehnung;
   //
         A     "DB1001_TT_State".Bits.Taktdehnung;
         AN    "DB1001_TT_State".IPOS.Status.RT_in_Position;
         A     "Flag_01_000_Hertz";
         O;
         A     "DB1001_TT_State".Bits.Taktdehnung;
         A     "DB1001_TT_State".IPOS.Status.RT_in_Position;
         A     "Flag_05_000_Hertz";
         O     "DB1001_TT_State".BA_Anlage.Lampentest;
         =     "LED_extend_cycle";
END_REGION

REGION Network 4: Freigabe zum Takten der Anlage

         AN    "DB1001_TT_State".Bits.Stop_fuer_WW;
         AN    "DB1001_TT_State".Bits.Stop_fuer_Teachen;
         AN    "DB1001_TT_State".Bits.StopAfterEmpty;

         AN    "DB005_RS<->Extern".MC_Interface[1].Data_from_MC.Shot_release;
         AN    "DB005_RS<->Extern".MC_Interface[1].Data_from_MC.Shot_preperation;
         AN    "DB1001_TT_State".BA_Anlage.Stop_angefordert;
         AN    "DB1030_TT_AddFaults".SafteyDeviceSelected[1];
         AN    "DB1030_TT_AddFaults".SafteyDeviceSelected[2];
         AN    "DB1030_TT_AddFaults".SafteyDeviceSelected[3];

         A     #Temp_Drehfreigabe;
         AN    "DB1001_TT_State".Bits.Taktdehnung;
         A     "DB1001_TT_State".BA_Anlage.Automatik;
         =     #Temp_Taktfreigabe;
END_REGION

REGION Network 5: Taktimpuls bilden
         CALL  "FC1041_TT_Taktimpuls"
         ( IN_Drehfreigabe         := #Temp_Taktfreigabe,
           IN_Taktfreigabe         := #Temp_Drehfreigabe,
           IN_Anlage_in_Position   := "DB1001_TT_State".IPOS.Status.RT_in_Position,
           IN_Start_Anlagenbetrieb := "DB1001_TT_State".BA_Anlage.Produktion,
           IN_Anlagenbetrieb       := "DB1001_TT_State".BA_Anlage.Start_Produktion,
           IN_DW_Taktzeit          := "DB1049_TT_Value".Taktzeit,
           IN_Takttimer            := "TMTT_Tact",
           IN_Vorwarnzeit_1_in_Dec := 5,
           IN_Vorwarnzeit_2_in_Dec := 3,
           IO_Status               := "DB1001_TT_State".Takt
         );
   //-----
END_REGION

REGION Network 6: Sollwerte an FU
         L     "DB1049_TT_Value".Antrieb_RP;
         T     #Temp_Rampe_Plus;
         L     "DB1049_TT_Value".Antrieb_RN;
         T     #Temp_Rampe_Minus;
         L     "DB1049_TT_Value".Antrieb_Hand;
         T     #Temp_Speed_Hand;
         L     "DB1049_TT_Value".Antrieb_Auto;
         T     #Temp_Speed_Automatik;
   //-----
         L     0;
         A     "DB1001_TT_State".Bits.Stop_fuer_WW;
         JCN   Off2;
         L     "DB1049_TT_Value".Pos_Offset_WW;
         JU    Off;
   Off2: NOP   0;
         A     "DB1001_TT_State".Bits.Stop_fuer_Teachen;
         JCN   Off3;
         L     "DB1049_TT_Value".Pos_Offset_Teachen;
         JU    Off;
   Off3: NOP   0;
   Off:  T     #Temp_Offset_Position;
END_REGION

REGION Network 7: Umrichter für Rundtisch ansteuern
         A     "Button_Tip_+";
         A     "DB1001_TT_State".BA_Anlage.Hand;
         =     "Button_Tip_+";

         A     "Button_Tip_-";
         A     "DB1001_TT_State".BA_Anlage.Hand;
         =     "Button_Tip_-";

   // Genauhalt INI
         L     "DB1001_TT_State".IPOS.Status.Aktuelle_Position;
         L     0;
         ==I;
         A     "DB1001_TT_State".IPOS.Eingaenge_von_IPOS.Ipos_referenziert;
         =     #Temp_GenauhalteSignal;
   //-----
         CALL  "FC1042_RT_IPOS_CTRL"
         ( IN_EA_Adresse            := 700,
           IN_Taktend               := TRUE,
           IN_Taktend_1_Segment     := TRUE,
           IN_DP_ok                 := TRUE,
           IN_IPOS_referenziert     := "DB1001_TT_State".IPOS.Eingaenge_von_IPOS.Ipos_referenziert,
           IN_Stoerung_Luefter      := FALSE,
           IN_Motorschutz           := "F_FC_turn_table",
           IN_STG_Umrichter         := "F_fuse_FC_turn_table",
           IN_Reset_fault_Fkt       := "DB1011_TT_Fault".Reset_FC_RT,
           IN_Kettenspanner_ok      := TRUE,
           IN_Drehsperre            := #Temp_Drehsperre,
           IN_HW_und_BA_ok          := "DB1001_TT_State".BA_Anlage.Aktiv,
           IN_AutoStop_ok           := "DB1001_TT_State".BA_Anlage.Automatik_Stop_ok,
           IN_BA_Hand               := "DB1001_TT_State".BA_Anlage.Hand,
           IN_BA_Automatik          := "DB1001_TT_State".BA_Anlage.Automatik,
           IN_BA_Referenzieren      := "DB1001_TT_State".BA_Anlage.Referenzieren,
           IN_BA_Start_Taktbetrieb  := "DB1001_TT_State".BA_Anlage.Start_Produktion,
           IN_BA_Taktbetrieb        := "DB1001_TT_State".BA_Anlage.Produktion,
           IN_BA_Stop_angefordert   := "DB1001_TT_State".BA_Anlage.Stop_angefordert,
           IN_BA_Lampentest         := "DB1001_TT_State".BA_Anlage.Lampentest,
           IN_Taktimpuls            := "DB1001_TT_State".Takt.Taktimpuls,
           IN_T_Tippen_plus         := "Button_Tip_+",
           IN_T_Tippen_minus        := "Button_Tip_-",
           IN_Genauhaltini          := #Temp_GenauhalteSignal,
           IN_Anzahl_Segmente       := #Temp_AmoutOfSegments,
           IN_DW_Rampe_Pos          := #Temp_Rampe_Plus,
           IN_DW_Rampe_Neg          := #Temp_Rampe_Minus,
           IN_DW_Speed_Hand         := #Temp_Speed_Hand,
           IN_DW_Speed_Automatik    := #Temp_Speed_Automatik,
           IN_DW_Offset_Position    := #Temp_Offset_Position,
           IN_TM_Universal          := "TMTT_IPOS_Universal",
           IN_TM_Freigabe           := "TMTT_IPOS_Enable",
           IN_TM_Tol_Genauhalt      := "TMTT_IPOS_TolInPos",
           IN_TM_Verz_STG_FU        := "TMTT_IPOS_FaultFC",
           IN_TM_Verz_Ziel_erreicht := "TMTT_IPOS_DelayInPos",
           IN_TM_AnfahrWarnung      := "TMTT_IPOS_Horn",
           IN_ZT_Tol_Genauhalt      := S5T#1S,
           IN_Time_Anfahrwarnung    := "DB1049_TT_Value".Vorwarnzeit,
           OUT_aktuelle_Position    := "DB1001_TT_State".Aktuelle_Position,
           OUT_FRG_Umrichter        := "Release_FC_turn_table",
           OUT_H_Tippen_plus        := "LED_Tip_+",
           OUT_H_Tippen_minus       := "LED_Tip_-",
           OUT_H_Referenzpunkt      := "LED_reference_TT",
           OUT_H_AnfahrWarnung      := #Temp_AnfahrWarnung,
           IO_Status                := "DB1001_TT_State".IPOS,
           IO_Fault                 := "DB1040_TT_MovementFault".IPOS,
           IO_New_Fault             := "DB1011_TT_Fault".Stoerungsaend_RT,
           IO_Fault_GRP_1           := "DB1011_TT_Fault".STG1_RT,
           IO_Fault_GRP_2           := "DB1011_TT_Fault".STG2_RT,
           IO_Fault_GRP_3           := "DB1011_TT_Fault".STG3_RT
         );
   //-----
END_REGION

REGION Network 8: Ansteuerung Vorwarnhupe
         O     "DB1001_TT_State".BA_Anlage.Anfahrwarnung;
   //      O     "DB1001_TT_State".Takt.Vorwarnung_1
         O     #Temp_AnfahrWarnung;
         =     "LED_start_cycle";
END_REGION

REGION Network 9: Positionsabhängige Freigaben bilden
   // Der Bereich eines Segmentes ist 18°.
   // Die eingegebenen Werte müssen zwischen 0 (0°) und 180 (18°) liegen.
         A     "DB1001_TT_State".IPOS.Status.RT_in_Position;
         A     "DB1001_TT_State".IPOS.Status.IPOS_referenziert;
         =     "DB1001_TT_State".Segment_in_Position.Reserve1;
   //
         A(;
         L     "DB1001_TT_State".Aktuelle_Position;
         L     10;
         >=D;
         );
         A(;
         L     "DB1001_TT_State".Aktuelle_Position;
         L     15;
         <D;
         );
         A     "DB1001_TT_State".IPOS.Status.IPOS_referenziert;
         =     "DB1001_TT_State".Segment_in_Position.FRG_abloeschen_Programm;
   //
         A(;
         L     "DB1001_TT_State".Aktuelle_Position;
         L     50;
         >=D;
         );
         A(;
         L     "DB1001_TT_State".Aktuelle_Position;
         L     55;
         <D;
         );
         A     "DB1001_TT_State".IPOS.Status.IPOS_referenziert;
         =     "DB1001_TT_State".Segment_in_Position.Reserve3;
   //
         A(;
         L     "DB1001_TT_State".Aktuelle_Position;
         L     5;
         >=D;
         );
         A(;
         L     "DB1001_TT_State".Aktuelle_Position;
         L     10;
         <D;
         );
         A     "DB1001_TT_State".IPOS.Status.IPOS_referenziert;
         =     "DB1001_TT_State".Segment_in_Position.Reserve5;
   //
         A(;
         L     "DB1001_TT_State".Aktuelle_Position;
         L     120;
         >=D;
         );
         A(;
         L     "DB1001_TT_State".Aktuelle_Position;
         L     125;
         <D;
         );
         A     "DB1001_TT_State".IPOS.Status.IPOS_referenziert;
         =     "DB1001_TT_State".Segment_in_Position.Test_IFM_Initiator;
   //
         A(;
         L     "DB1001_TT_State".Aktuelle_Position;
         L     140;
         >=D;
         );
         A(;
         L     "DB1001_TT_State".Aktuelle_Position;
         L     145;
         <D;
         );
         A     "DB1001_TT_State".IPOS.Status.IPOS_referenziert;
         =     "DB1001_TT_State".Segment_in_Position.Start_Schaeumen;
   //
         A     "DB1001_TT_State".IPOS.Status.IPOS_referenziert;
         A     "DB1001_TT_State".IPOS.Status.RT_in_Position;
         =     "DB1001_TT_State".Segment_in_Position.FRG_Schaeumen;
END_REGION

REGION Network 10: Segmentkennung
         CALL  "FC1045_getStationRW"
         ( Anzahl_Segmente := #Temp_AmoutOfSegments,
           Maxwert         := 3600,
           Offset          := 50,
           Istwert         := "DB1001_TT_State".IPOS.Eingaenge_von_IPOS.Istposition,
           SegmenteReverse := FALSE,
           Ret_Val         := "DB1001_TT_State".Segmentkennung.Seg_No_Stat_1
         );
   //---
         A     "DB1001_TT_State".IPOS.Status.IPOS_referenziert;
         JC    Tran;
         L     0;
         T     "DB1001_TT_State".Segmentkennung.Seg_No_Stat_1;
   Tran: NOP   0;
END_REGION

REGION Network 11: Stationsbelegung
         CALL  "FC1046_SegmInStation"
         ( IN_Amount_Segment := #Temp_AmoutOfSegments
         );
END_REGION
END_FUNCTION

